REGION Network 13: DB60 DBX2.0 = FS332 No Flow
   // GCU_ALARM_WORD_02_BIT_0
   RUNG wire#powerrail
      Contact( "300_AUT_SEQ_TMRS_DB"."FS332 Delay".Q )
      { S7_Templates := "SrcType := Int" } GE_Contact(in1 := "100_GCU_AUTO_SEQ_DB".CRNT_STEP, in2 := 60)
      { S7_Templates := "SrcType := Int" } LE_Contact(in1 := "100_GCU_AUTO_SEQ_DB".CRNT_STEP, in2 := 560)
      S_Coil( %DB60.DBX2.0 )
   END_RUNG
   // the same network as SCL:
   IF "300_AUT_SEQ_TMRS_DB"."FS332 Delay".Q AND ("100_GCU_AUTO_SEQ_DB".CRNT_STEP >= 60) AND ("100_GCU_AUTO_SEQ_DB".CRNT_STEP <= 560) THEN
       %DB60.DBX2.0 := TRUE;
   END_IF;
END_REGION

REGION Network 14: DB60 DBX2.1 = PIT348 LOLO
   // GCU_ALARM_WORD_02_BIT_1      changed to 60 to 120 for test
   RUNG wire#powerrail
      { S7_Templates := "SrcType := Int" } GE_Contact(in1 := "100_GCU_AUTO_SEQ_DB".CRNT_STEP, in2 := 140)
      { S7_Templates := "SrcType := Int" } LT_Contact(in1 := "100_GCU_AUTO_SEQ_DB".CRNT_STEP, in2 := 540)
      Contact( "PIT348_ALM_ANALOG_DB73"."ALARM LL" )
      I_Contact( "10_DI_DATA"."FS_332 FLW_OK" )
      S_Coil( %DB60.DBX2.1 )
   END_RUNG
   // the same network as SCL:
   IF ("100_GCU_AUTO_SEQ_DB".CRNT_STEP >= 140) AND ("100_GCU_AUTO_SEQ_DB".CRNT_STEP < 540) AND "PIT348_ALM_ANALOG_DB73"."ALARM LL" AND NOT "10_DI_DATA"."FS_332 FLW_OK" THEN
       %DB60.DBX2.1 := TRUE;
   END_IF;
END_REGION

REGION Network 15: DB60 DBX2.2 = PIT348 HIHI
   // GCU_ALARM_WORD_02_BIT_2
   RUNG wire#powerrail
      Contact( "PIT348_ALM_ANALOG_DB73"."ALARM HH" )
      I_Contact( "10_DI_DATA"."FS_332 FLW_OK" )
      S_Coil( %DB60.DBX2.2 )
   END_RUNG
   // the same network as SCL:
   IF "PIT348_ALM_ANALOG_DB73"."ALARM HH" AND NOT "10_DI_DATA"."FS_332 FLW_OK" THEN
       %DB60.DBX2.2 := TRUE;
   END_IF;
END_REGION

REGION Network 16: DB60 DBX2.3 = FS350 Low Flow
   // GCU_ALARM_WORD_02_BIT_3
   RUNG wire#powerrail
      Contact( "TIT406_ALM_ANALOG_DB74".Error_present )
      Contact( "TIT408_ALM_ANALOG_DB75".Error_present )
      I_Contact( "10_DI_DATA".FS_350_FLW_OK )
      S_Coil( %DB60.DBX2.3 )
   END_RUNG
   // the same network as SCL:
   IF "TIT406_ALM_ANALOG_DB74".Error_present AND "TIT408_ALM_ANALOG_DB75".Error_present AND NOT "10_DI_DATA".FS_350_FLW_OK THEN
       %DB60.DBX2.3 := TRUE;
   END_IF;
END_REGION

REGION Network 17: DB60 DBX2.5 = TT002 HIHI
   // GCU_ALARM_WORD_02_BIT_5
   RUNG wire#powerrail
      Contact( "TT002_ALM_ANALOG_DB76"."ALARM HH" )
      S_Coil( %DB60.DBX2.5 )
   END_RUNG
   // the same network as SCL:
   IF "TT002_ALM_ANALOG_DB76"."ALARM HH" THEN %DB60.DBX2.5 := TRUE; END_IF;
END_REGION

REGION Network 18: DB60 DBX2.6 = PT002 HIHI
   // GCU_ALARM_WORD_02_BIT_6
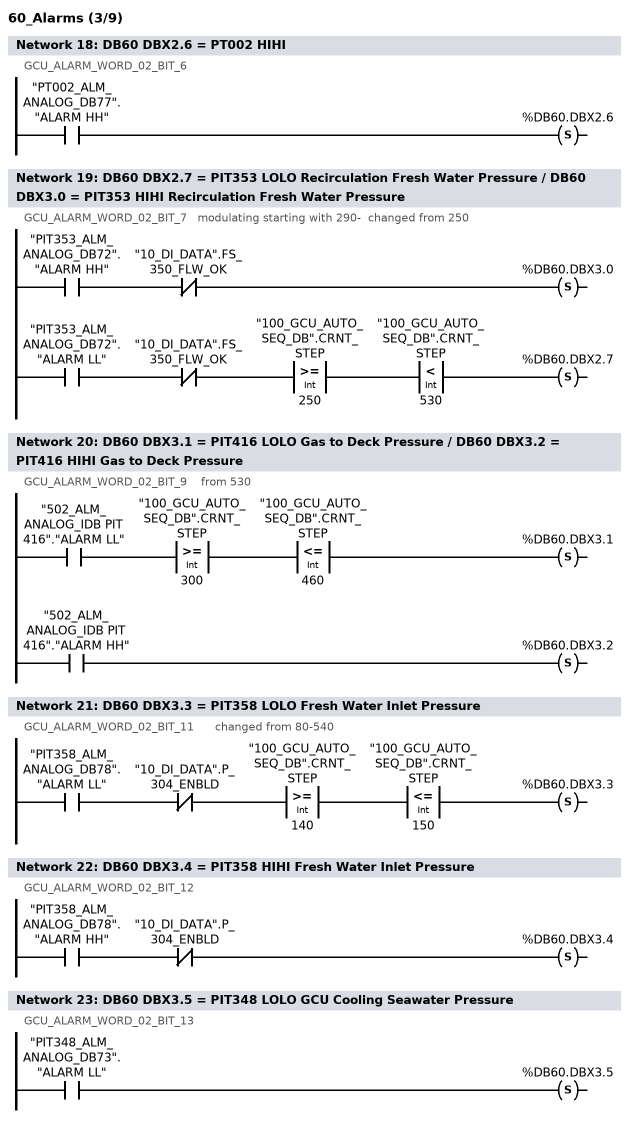
   RUNG wire#powerrail
      Contact( "PT002_ALM_ANALOG_DB77"."ALARM HH" )
      S_Coil( %DB60.DBX2.6 )
   END_RUNG
   // the same network as SCL:
   IF "PT002_ALM_ANALOG_DB77"."ALARM HH" THEN %DB60.DBX2.6 := TRUE; END_IF;
END_REGION

REGION Network 19: DB60 DBX2.7 = PIT353 LOLO Recirculation Fresh Water Pressure / DB60 DBX3.0 = PIT353 HIHI Recirculation Fresh Water Pressure
   // GCU_ALARM_WORD_02_BIT_7   modulating starting with 290-  changed from 250
   RUNG wire#powerrail
      Contact( "PIT353_ALM_ANALOG_DB72"."ALARM HH" )
      I_Contact( "10_DI_DATA".FS_350_FLW_OK )
      S_Coil( %DB60.DBX3.0 )
   END_RUNG
   RUNG wire#powerrail
      Contact( "PIT353_ALM_ANALOG_DB72"."ALARM LL" )
      I_Contact( "10_DI_DATA".FS_350_FLW_OK )
      { S7_Templates := "SrcType := Int" } GE_Contact(in1 := "100_GCU_AUTO_SEQ_DB".CRNT_STEP, in2 := 250)
      { S7_Templates := "SrcType := Int" } LT_Contact(in1 := "100_GCU_AUTO_SEQ_DB".CRNT_STEP, in2 := 530)
      S_Coil( %DB60.DBX2.7 )
   END_RUNG
   // the same network as SCL:
   IF "PIT353_ALM_ANALOG_DB72"."ALARM HH" AND NOT "10_DI_DATA".FS_350_FLW_OK THEN
       %DB60.DBX3.0 := TRUE;
   END_IF;
   IF "PIT353_ALM_ANALOG_DB72"."ALARM LL" AND NOT "10_DI_DATA".FS_350_FLW_OK AND ("100_GCU_AUTO_SEQ_DB".CRNT_STEP >= 250) AND ("100_GCU_AUTO_SEQ_DB".CRNT_STEP < 530) THEN
       %DB60.DBX2.7 := TRUE;
   END_IF;
END_REGION

REGION Network 20: DB60 DBX3.1 = PIT416 LOLO Gas to Deck Pressure / DB60 DBX3.2 = PIT416 HIHI Gas to Deck Pressure
   // GCU_ALARM_WORD_02_BIT_9    from 530
   RUNG wire#powerrail
      Contact( "502_ALM_ANALOG_IDB PIT 416"."ALARM LL" )
      { S7_Templates := "SrcType := Int" } GE_Contact(in1 := "100_GCU_AUTO_SEQ_DB".CRNT_STEP, in2 := 300)
      { S7_Templates := "SrcType := Int" } LE_Contact(in1 := "100_GCU_AUTO_SEQ_DB".CRNT_STEP, in2 := 460)
      S_Coil( %DB60.DBX3.1 )
   END_RUNG
   RUNG wire#powerrail
      Contact( "502_ALM_ANALOG_IDB PIT 416"."ALARM HH" )
      S_Coil( %DB60.DBX3.2 )
   END_RUNG
   // the same network as SCL:
   IF "502_ALM_ANALOG_IDB PIT 416"."ALARM LL" AND ("100_GCU_AUTO_SEQ_DB".CRNT_STEP >= 300) AND ("100_GCU_AUTO_SEQ_DB".CRNT_STEP <= 460) THEN
       %DB60.DBX3.1 := TRUE;
   END_IF;
   IF "502_ALM_ANALOG_IDB PIT 416"."ALARM HH" THEN %DB60.DBX3.2 := TRUE; END_IF;
END_REGION

REGION Network 21: DB60 DBX3.3 = PIT358 LOLO Fresh Water Inlet Pressure
   // GCU_ALARM_WORD_02_BIT_11      changed from 80-540
   RUNG wire#powerrail
      Contact( "PIT358_ALM_ANALOG_DB78"."ALARM LL" )
      I_Contact( "10_DI_DATA".P_304_ENBLD )
      { S7_Templates := "SrcType := Int" } GE_Contact(in1 := "100_GCU_AUTO_SEQ_DB".CRNT_STEP, in2 := 140)
      { S7_Templates := "SrcType := Int" } LE_Contact(in1 := "100_GCU_AUTO_SEQ_DB".CRNT_STEP, in2 := 150)
      S_Coil( %DB60.DBX3.3 )
   END_RUNG
   // the same network as SCL:
   IF "PIT358_ALM_ANALOG_DB78"."ALARM LL" AND NOT "10_DI_DATA".P_304_ENBLD AND ("100_GCU_AUTO_SEQ_DB".CRNT_STEP >= 140) AND ("100_GCU_AUTO_SEQ_DB".CRNT_STEP <= 150) THEN
       %DB60.DBX3.3 := TRUE;
   END_IF;
END_REGION

REGION Network 22: DB60 DBX3.4 = PIT358 HIHI Fresh Water Inlet Pressure
   // GCU_ALARM_WORD_02_BIT_12
   RUNG wire#powerrail
      Contact( "PIT358_ALM_ANALOG_DB78"."ALARM HH" )
      I_Contact( "10_DI_DATA".P_304_ENBLD )
      S_Coil( %DB60.DBX3.4 )
   END_RUNG
   // the same network as SCL:
   IF "PIT358_ALM_ANALOG_DB78"."ALARM HH" AND NOT "10_DI_DATA".P_304_ENBLD THEN %DB60.DBX3.4 := TRUE; END_IF;
END_REGION

REGION Network 23: DB60 DBX3.5 = PIT348 LOLO GCU Cooling Seawater Pressure
   // GCU_ALARM_WORD_02_BIT_13
   RUNG wire#powerrail
      Contact( "PIT348_ALM_ANALOG_DB73"."ALARM LL" )
      S_Coil( %DB60.DBX3.5 )
   END_RUNG
   // the same network as SCL:
   IF "PIT348_ALM_ANALOG_DB73"."ALARM LL" THEN %DB60.DBX3.5 := TRUE; END_IF;
END_REGION

REGION Network 24: DB60 DBX3.6 = PIT348 HIHI GCU Cooling Seawater Pressure
   // GCU_ALARM_WORD_02_BIT_14
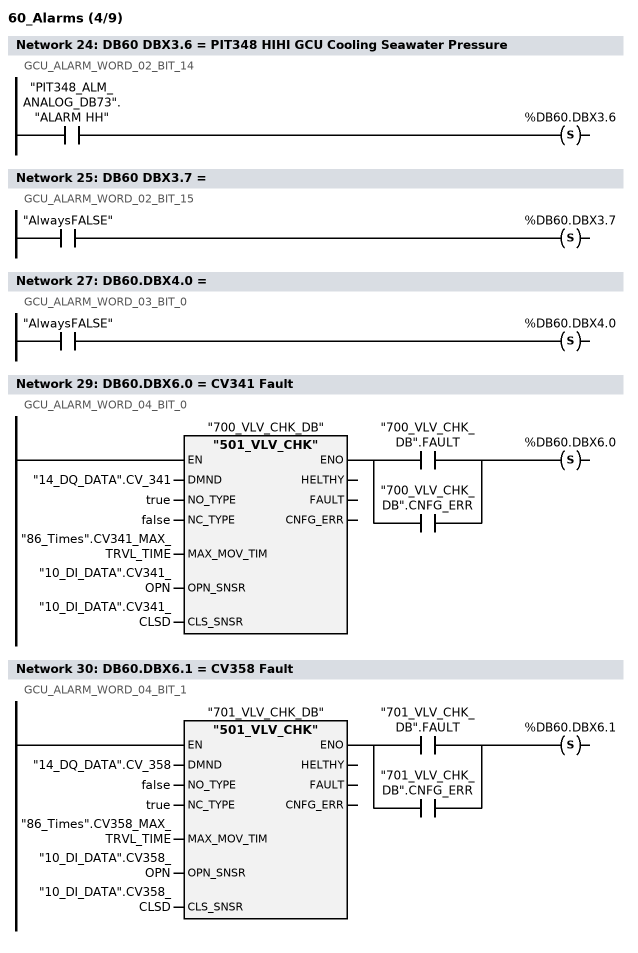
   RUNG wire#powerrail
      Contact( "PIT348_ALM_ANALOG_DB73"."ALARM HH" )
      S_Coil( %DB60.DBX3.6 )
   END_RUNG
   // the same network as SCL:
   IF "PIT348_ALM_ANALOG_DB73"."ALARM HH" THEN %DB60.DBX3.6 := TRUE; END_IF;
END_REGION

REGION Network 25: DB60 DBX3.7 =
   // GCU_ALARM_WORD_02_BIT_15
   RUNG wire#powerrail
      Contact( "AlwaysFALSE" )
      S_Coil( %DB60.DBX3.7 )
   END_RUNG
   // the same network as SCL:
   IF "AlwaysFALSE" THEN %DB60.DBX3.7 := TRUE; END_IF;
END_REGION

REGION Network 27: DB60.DBX4.0 =
   // GCU_ALARM_WORD_03_BIT_0
   RUNG wire#powerrail
      Contact( "AlwaysFALSE" )
      S_Coil( %DB60.DBX4.0 )
   END_RUNG
   // the same network as SCL:
   IF "AlwaysFALSE" THEN %DB60.DBX4.0 := TRUE; END_IF;
END_REGION

REGION Network 29: DB60.DBX6.0 = CV341 Fault
   // GCU_ALARM_WORD_04_BIT_0
   RUNG wire#powerrail
      "700_VLV_CHK_DB"(DMND := "14_DQ_DATA".CV_341, NO_TYPE := true, NC_TYPE := false, MAX_MOV_TIM := "86_Times".CV341_MAX_TRVL_TIME, OPN_SNSR := "10_DI_DATA".CV341_OPN, CLS_SNSR := "10_DI_DATA".CV341_CLSD, HELTHY =>, FAULT =>, CNFG_ERR =>)
      wire#w1
      Contact( "700_VLV_CHK_DB".FAULT )
      wire#w2
      S_Coil( %DB60.DBX6.0 )
   END_RUNG
   RUNG wire#w1
      Contact( "700_VLV_CHK_DB".CNFG_ERR )
   END_RUNG wire#w2
   // the same network as SCL:
   "700_VLV_CHK_DB"(DMND := "14_DQ_DATA".CV_341,   // "501_VLV_CHK"
                    NO_TYPE := true,
                    NC_TYPE := false,
                    MAX_MOV_TIM := "86_Times".CV341_MAX_TRVL_TIME,
                    OPN_SNSR := "10_DI_DATA".CV341_OPN,
                    CLS_SNSR := "10_DI_DATA".CV341_CLSD,
                    ENO => #_w1);
   IF #_w1 AND ("700_VLV_CHK_DB".FAULT OR "700_VLV_CHK_DB".CNFG_ERR) THEN %DB60.DBX6.0 := TRUE; END_IF;
END_REGION

REGION Network 30: DB60.DBX6.1 = CV358 Fault
   // GCU_ALARM_WORD_04_BIT_1
   RUNG wire#powerrail
      "701_VLV_CHK_DB"(DMND := "14_DQ_DATA".CV_358, NO_TYPE := false, NC_TYPE := true, MAX_MOV_TIM := "86_Times".CV358_MAX_TRVL_TIME, OPN_SNSR := "10_DI_DATA".CV358_OPN, CLS_SNSR := "10_DI_DATA".CV358_CLSD, HELTHY =>, FAULT =>, CNFG_ERR =>)
      wire#w1
      Contact( "701_VLV_CHK_DB".FAULT )
      wire#w2
      S_Coil( %DB60.DBX6.1 )
   END_RUNG
   RUNG wire#w1
      Contact( "701_VLV_CHK_DB".CNFG_ERR )
   END_RUNG wire#w2
   // the same network as SCL:
   "701_VLV_CHK_DB"(DMND := "14_DQ_DATA".CV_358,   // "501_VLV_CHK"
                    NO_TYPE := false,
                    NC_TYPE := true,
                    MAX_MOV_TIM := "86_Times".CV358_MAX_TRVL_TIME,
                    OPN_SNSR := "10_DI_DATA".CV358_OPN,
                    CLS_SNSR := "10_DI_DATA".CV358_CLSD,
                    ENO => #_w1);
   IF #_w1 AND ("701_VLV_CHK_DB".FAULT OR "701_VLV_CHK_DB".CNFG_ERR) THEN %DB60.DBX6.1 := TRUE; END_IF;
END_REGION

REGION Network 31: DB60.DBX6.2 = CV406 Fault
   // GCU_ALARM_WORD_04_BIT_2
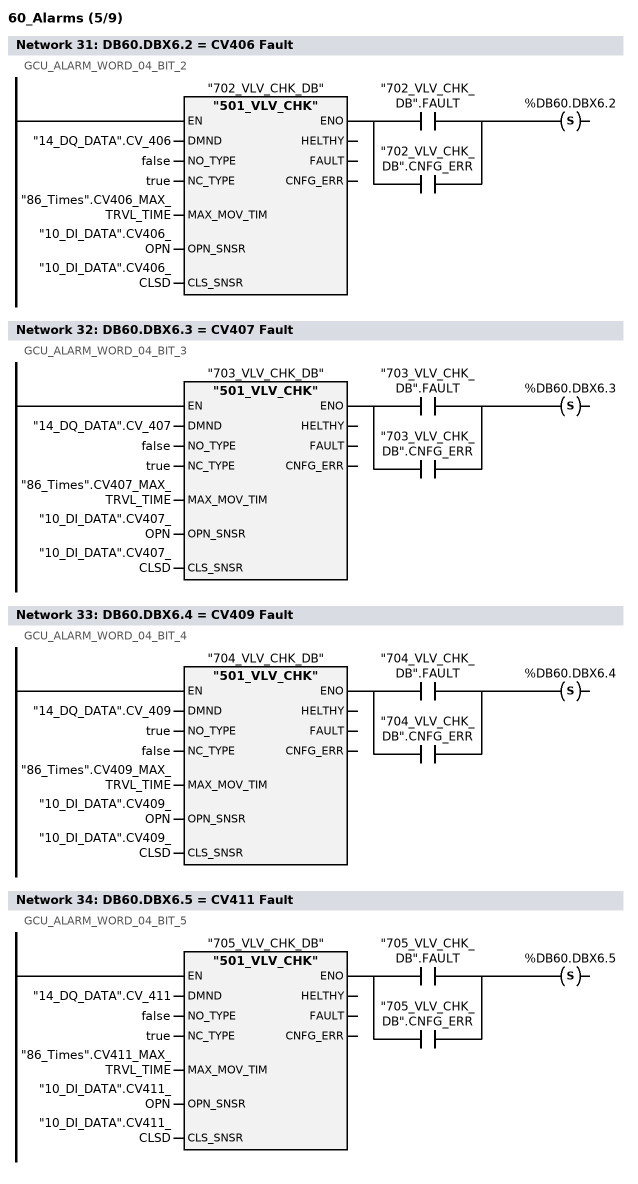
   RUNG wire#powerrail
      "702_VLV_CHK_DB"(DMND := "14_DQ_DATA".CV_406, NO_TYPE := false, NC_TYPE := true, MAX_MOV_TIM := "86_Times".CV406_MAX_TRVL_TIME, OPN_SNSR := "10_DI_DATA".CV406_OPN, CLS_SNSR := "10_DI_DATA".CV406_CLSD, HELTHY =>, FAULT =>, CNFG_ERR =>)
      wire#w1
      Contact( "702_VLV_CHK_DB".FAULT )
      wire#w2
      S_Coil( %DB60.DBX6.2 )
   END_RUNG
   RUNG wire#w1
      Contact( "702_VLV_CHK_DB".CNFG_ERR )
   END_RUNG wire#w2
   // the same network as SCL:
   "702_VLV_CHK_DB"(DMND := "14_DQ_DATA".CV_406,   // "501_VLV_CHK"
                    NO_TYPE := false,
                    NC_TYPE := true,
                    MAX_MOV_TIM := "86_Times".CV406_MAX_TRVL_TIME,
                    OPN_SNSR := "10_DI_DATA".CV406_OPN,
                    CLS_SNSR := "10_DI_DATA".CV406_CLSD,
                    ENO => #_w1);
   IF #_w1 AND ("702_VLV_CHK_DB".FAULT OR "702_VLV_CHK_DB".CNFG_ERR) THEN %DB60.DBX6.2 := TRUE; END_IF;
END_REGION

REGION Network 32: DB60.DBX6.3 = CV407 Fault
   // GCU_ALARM_WORD_04_BIT_3
   RUNG wire#powerrail
      "703_VLV_CHK_DB"(DMND := "14_DQ_DATA".CV_407, NO_TYPE := false, NC_TYPE := true, MAX_MOV_TIM := "86_Times".CV407_MAX_TRVL_TIME, OPN_SNSR := "10_DI_DATA".CV407_OPN, CLS_SNSR := "10_DI_DATA".CV407_CLSD, HELTHY =>, FAULT =>, CNFG_ERR =>)
      wire#w1
      Contact( "703_VLV_CHK_DB".FAULT )
      wire#w2
      S_Coil( %DB60.DBX6.3 )
   END_RUNG
   RUNG wire#w1
      Contact( "703_VLV_CHK_DB".CNFG_ERR )
   END_RUNG wire#w2
   // the same network as SCL:
   "703_VLV_CHK_DB"(DMND := "14_DQ_DATA".CV_407,   // "501_VLV_CHK"
                    NO_TYPE := false,
                    NC_TYPE := true,
                    MAX_MOV_TIM := "86_Times".CV407_MAX_TRVL_TIME,
                    OPN_SNSR := "10_DI_DATA".CV407_OPN,
                    CLS_SNSR := "10_DI_DATA".CV407_CLSD,
                    ENO => #_w1);
   IF #_w1 AND ("703_VLV_CHK_DB".FAULT OR "703_VLV_CHK_DB".CNFG_ERR) THEN %DB60.DBX6.3 := TRUE; END_IF;
END_REGION

REGION Network 33: DB60.DBX6.4 = CV409 Fault
   // GCU_ALARM_WORD_04_BIT_4
   RUNG wire#powerrail
      "704_VLV_CHK_DB"(DMND := "14_DQ_DATA".CV_409, NO_TYPE := true, NC_TYPE := false, MAX_MOV_TIM := "86_Times".CV409_MAX_TRVL_TIME, OPN_SNSR := "10_DI_DATA".CV409_OPN, CLS_SNSR := "10_DI_DATA".CV409_CLSD, HELTHY =>, FAULT =>, CNFG_ERR =>)
      wire#w1
      Contact( "704_VLV_CHK_DB".FAULT )
      wire#w2
      S_Coil( %DB60.DBX6.4 )
   END_RUNG
   RUNG wire#w1
      Contact( "704_VLV_CHK_DB".CNFG_ERR )
   END_RUNG wire#w2
   // the same network as SCL:
   "704_VLV_CHK_DB"(DMND := "14_DQ_DATA".CV_409,   // "501_VLV_CHK"
                    NO_TYPE := true,
                    NC_TYPE := false,
                    MAX_MOV_TIM := "86_Times".CV409_MAX_TRVL_TIME,
                    OPN_SNSR := "10_DI_DATA".CV409_OPN,
                    CLS_SNSR := "10_DI_DATA".CV409_CLSD,
                    ENO => #_w1);
   IF #_w1 AND ("704_VLV_CHK_DB".FAULT OR "704_VLV_CHK_DB".CNFG_ERR) THEN %DB60.DBX6.4 := TRUE; END_IF;
END_REGION

REGION Network 34: DB60.DBX6.5 = CV411 Fault
   // GCU_ALARM_WORD_04_BIT_5
   RUNG wire#powerrail
      "705_VLV_CHK_DB"(DMND := "14_DQ_DATA".CV_411, NO_TYPE := false, NC_TYPE := true, MAX_MOV_TIM := "86_Times".CV411_MAX_TRVL_TIME, OPN_SNSR := "10_DI_DATA".CV411_OPN, CLS_SNSR := "10_DI_DATA".CV411_CLSD, HELTHY =>, FAULT =>, CNFG_ERR =>)
      wire#w1
      Contact( "705_VLV_CHK_DB".FAULT )
      wire#w2
      S_Coil( %DB60.DBX6.5 )
   END_RUNG
   RUNG wire#w1
      Contact( "705_VLV_CHK_DB".CNFG_ERR )
   END_RUNG wire#w2
   // the same network as SCL:
   "705_VLV_CHK_DB"(DMND := "14_DQ_DATA".CV_411,   // "501_VLV_CHK"
                    NO_TYPE := false,
                    NC_TYPE := true,
                    MAX_MOV_TIM := "86_Times".CV411_MAX_TRVL_TIME,
                    OPN_SNSR := "10_DI_DATA".CV411_OPN,
                    CLS_SNSR := "10_DI_DATA".CV411_CLSD,
                    ENO => #_w1);
   IF #_w1 AND ("705_VLV_CHK_DB".FAULT OR "705_VLV_CHK_DB".CNFG_ERR) THEN %DB60.DBX6.5 := TRUE; END_IF;
END_REGION

REGION Network 35: DB60.DBX6.6 = CV441 Fault
   // GCU_ALARM_WORD_04_BIT_6
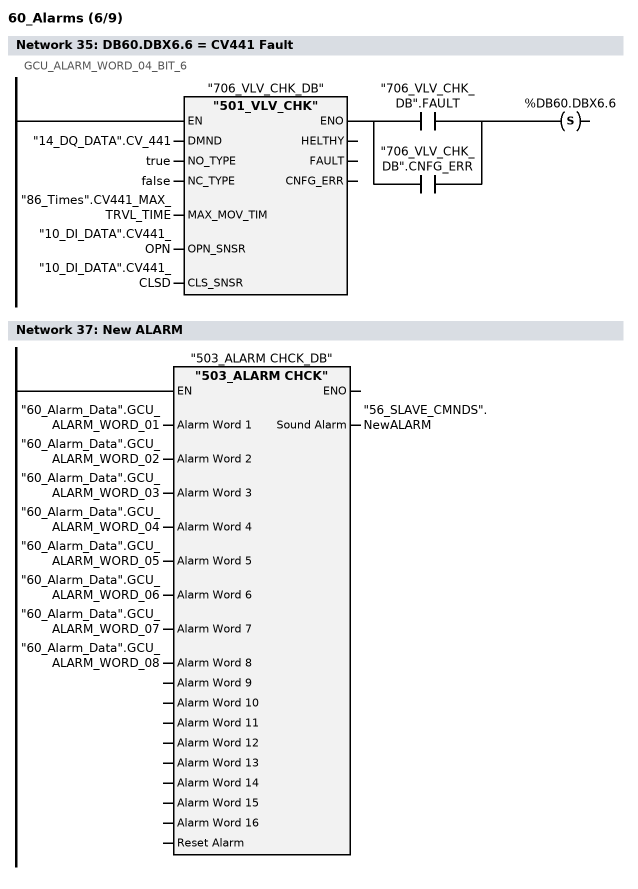
   RUNG wire#powerrail
      "706_VLV_CHK_DB"(DMND := "14_DQ_DATA".CV_441, NO_TYPE := true, NC_TYPE := false, MAX_MOV_TIM := "86_Times".CV441_MAX_TRVL_TIME, OPN_SNSR := "10_DI_DATA".CV441_OPN, CLS_SNSR := "10_DI_DATA".CV441_CLSD, HELTHY =>, FAULT =>, CNFG_ERR =>)
      wire#w1
      Contact( "706_VLV_CHK_DB".FAULT )
      wire#w2
      S_Coil( %DB60.DBX6.6 )
   END_RUNG
   RUNG wire#w1
      Contact( "706_VLV_CHK_DB".CNFG_ERR )
   END_RUNG wire#w2
   // the same network as SCL:
   "706_VLV_CHK_DB"(DMND := "14_DQ_DATA".CV_441,   // "501_VLV_CHK"
                    NO_TYPE := true,
                    NC_TYPE := false,
                    MAX_MOV_TIM := "86_Times".CV441_MAX_TRVL_TIME,
                    OPN_SNSR := "10_DI_DATA".CV441_OPN,
                    CLS_SNSR := "10_DI_DATA".CV441_CLSD,
                    ENO => #_w1);
   IF #_w1 AND ("706_VLV_CHK_DB".FAULT OR "706_VLV_CHK_DB".CNFG_ERR) THEN %DB60.DBX6.6 := TRUE; END_IF;
END_REGION

REGION Network 37: New ALARM
   RUNG wire#powerrail
      "503_ALARM CHCK_DB"("Alarm Word 1" := "60_Alarm_Data".GCU_ALARM_WORD_01, "Alarm Word 2" := "60_Alarm_Data".GCU_ALARM_WORD_02, "Alarm Word 3" := "60_Alarm_Data".GCU_ALARM_WORD_03, "Alarm Word 4" := "60_Alarm_Data".GCU_ALARM_WORD_04, "Alarm Word 5" := "60_Alarm_Data".GCU_ALARM_WORD_05, "Alarm Word 6" := "60_Alarm_Data".GCU_ALARM_WORD_06, "Alarm Word 7" := "60_Alarm_Data".GCU_ALARM_WORD_07, "Alarm Word 8" := "60_Alarm_Data".GCU_ALARM_WORD_08, "Alarm Word 9" :=, "Alarm Word 10" :=, "Alarm Word 11" :=, "Alarm Word 12" :=, "Alarm Word 13" :=, "Alarm Word 14" :=, "Alarm Word 15" :=, "Alarm Word 16" :=, "Reset Alarm" :=, "Sound Alarm" => "56_SLAVE_CMNDS".NewALARM)
   END_RUNG
   // the same network as SCL:
   "503_ALARM CHCK_DB"("Alarm Word 1" := "60_Alarm_Data".GCU_ALARM_WORD_01,   // "503_ALARM CHCK"
                       "Alarm Word 2" := "60_Alarm_Data".GCU_ALARM_WORD_02,
                       "Alarm Word 3" := "60_Alarm_Data".GCU_ALARM_WORD_03,
                       "Alarm Word 4" := "60_Alarm_Data".GCU_ALARM_WORD_04,
                       "Alarm Word 5" := "60_Alarm_Data".GCU_ALARM_WORD_05,
                       "Alarm Word 6" := "60_Alarm_Data".GCU_ALARM_WORD_06,
                       "Alarm Word 7" := "60_Alarm_Data".GCU_ALARM_WORD_07,
                       "Alarm Word 8" := "60_Alarm_Data".GCU_ALARM_WORD_08,
                       "Sound Alarm" => "56_SLAVE_CMNDS".NewALARM);
END_REGION

REGION Network 38: Alarm Present
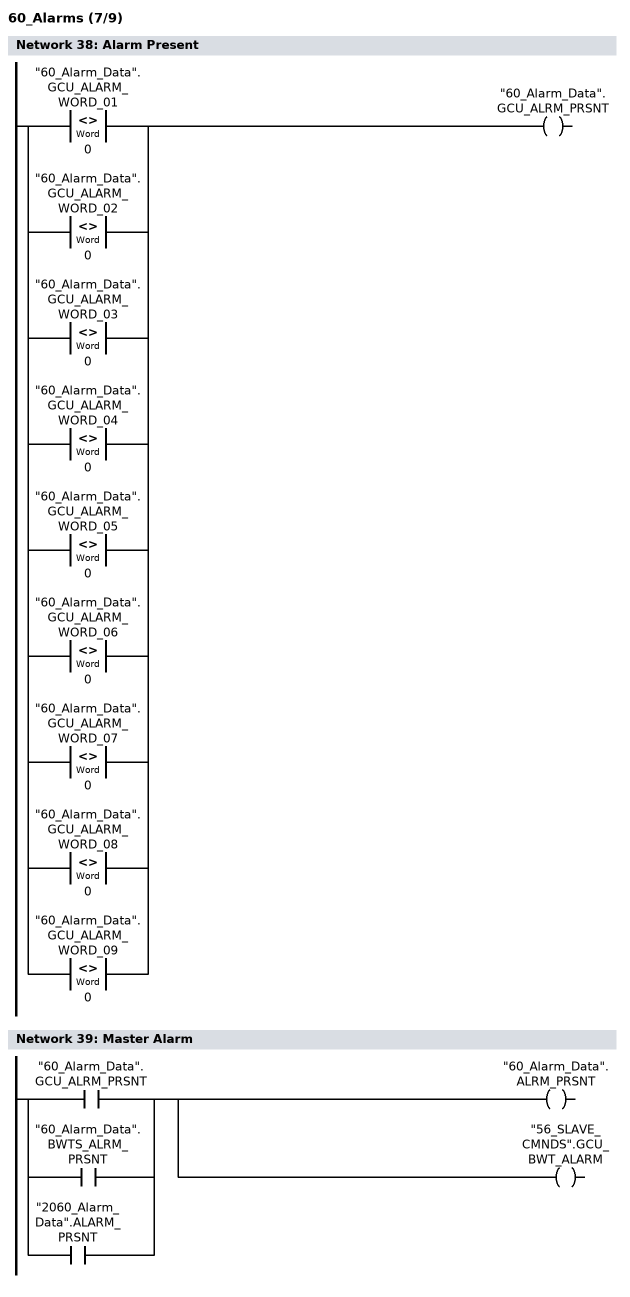
   RUNG wire#powerrail
      { S7_Templates := "SrcType := Word" } NE_Contact(in1 := "60_Alarm_Data".GCU_ALARM_WORD_01, in2 := 0)
      wire#w1
      Coil( "60_Alarm_Data".GCU_ALRM_PRSNT )
   END_RUNG
   RUNG wire#powerrail
      { S7_Templates := "SrcType := Word" } NE_Contact(in1 := "60_Alarm_Data".GCU_ALARM_WORD_02, in2 := 0)
   END_RUNG wire#w1
   RUNG wire#powerrail
      { S7_Templates := "SrcType := Word" } NE_Contact(in1 := "60_Alarm_Data".GCU_ALARM_WORD_03, in2 := 0)
   END_RUNG wire#w1
   RUNG wire#powerrail
      { S7_Templates := "SrcType := Word" } NE_Contact(in1 := "60_Alarm_Data".GCU_ALARM_WORD_04, in2 := 0)
   END_RUNG wire#w1
   RUNG wire#powerrail
      { S7_Templates := "SrcType := Word" } NE_Contact(in1 := "60_Alarm_Data".GCU_ALARM_WORD_05, in2 := 0)
   END_RUNG wire#w1
   RUNG wire#powerrail
      { S7_Templates := "SrcType := Word" } NE_Contact(in1 := "60_Alarm_Data".GCU_ALARM_WORD_06, in2 := 0)
   END_RUNG wire#w1
   RUNG wire#powerrail
      { S7_Templates := "SrcType := Word" } NE_Contact(in1 := "60_Alarm_Data".GCU_ALARM_WORD_07, in2 := 0)
   END_RUNG wire#w1
   RUNG wire#powerrail
      { S7_Templates := "SrcType := Word" } NE_Contact(in1 := "60_Alarm_Data".GCU_ALARM_WORD_08, in2 := 0)
   END_RUNG wire#w1
   RUNG wire#powerrail
      { S7_Templates := "SrcType := Word" } NE_Contact(in1 := "60_Alarm_Data".GCU_ALARM_WORD_09, in2 := 0)
   END_RUNG wire#w1
   // the same network as SCL:
   "60_Alarm_Data".GCU_ALRM_PRSNT := ("60_Alarm_Data".GCU_ALARM_WORD_01 <> 0) OR ("60_Alarm_Data".GCU_ALARM_WORD_02 <> 0) OR ("60_Alarm_Data".GCU_ALARM_WORD_03 <> 0) OR ("60_Alarm_Data".GCU_ALARM_WORD_04 <> 0) OR ("60_Alarm_Data".GCU_ALARM_WORD_05 <> 0) OR ("60_Alarm_Data".GCU_ALARM_WORD_06 <> 0) OR ("60_Alarm_Data".GCU_ALARM_WORD_07 <> 0) OR ("60_Alarm_Data".GCU_ALARM_WORD_08 <> 0) OR ("60_Alarm_Data".GCU_ALARM_WORD_09 <> 0);
END_REGION

REGION Network 39: Master Alarm
   RUNG wire#powerrail
      Contact( "60_Alarm_Data".GCU_ALRM_PRSNT )
      wire#w1
      Coil( "60_Alarm_Data".ALRM_PRSNT )
   END_RUNG
   RUNG wire#powerrail
      Contact( "60_Alarm_Data".BWTS_ALRM_PRSNT )
   END_RUNG wire#w1
   RUNG wire#powerrail
      Contact( "2060_Alarm_Data".ALARM_PRSNT )
   END_RUNG wire#w1
   RUNG wire#w1
      Coil( "56_SLAVE_CMNDS".GCU_BWT_ALARM )
   END_RUNG
   // the same network as SCL:
   "60_Alarm_Data".ALRM_PRSNT := "60_Alarm_Data".GCU_ALRM_PRSNT OR "60_Alarm_Data".BWTS_ALRM_PRSNT OR "2060_Alarm_Data".ALARM_PRSNT;
   "56_SLAVE_CMNDS".GCU_BWT_ALARM := "60_Alarm_Data".ALRM_PRSNT;
END_REGION

REGION Network 40: Alarm reset
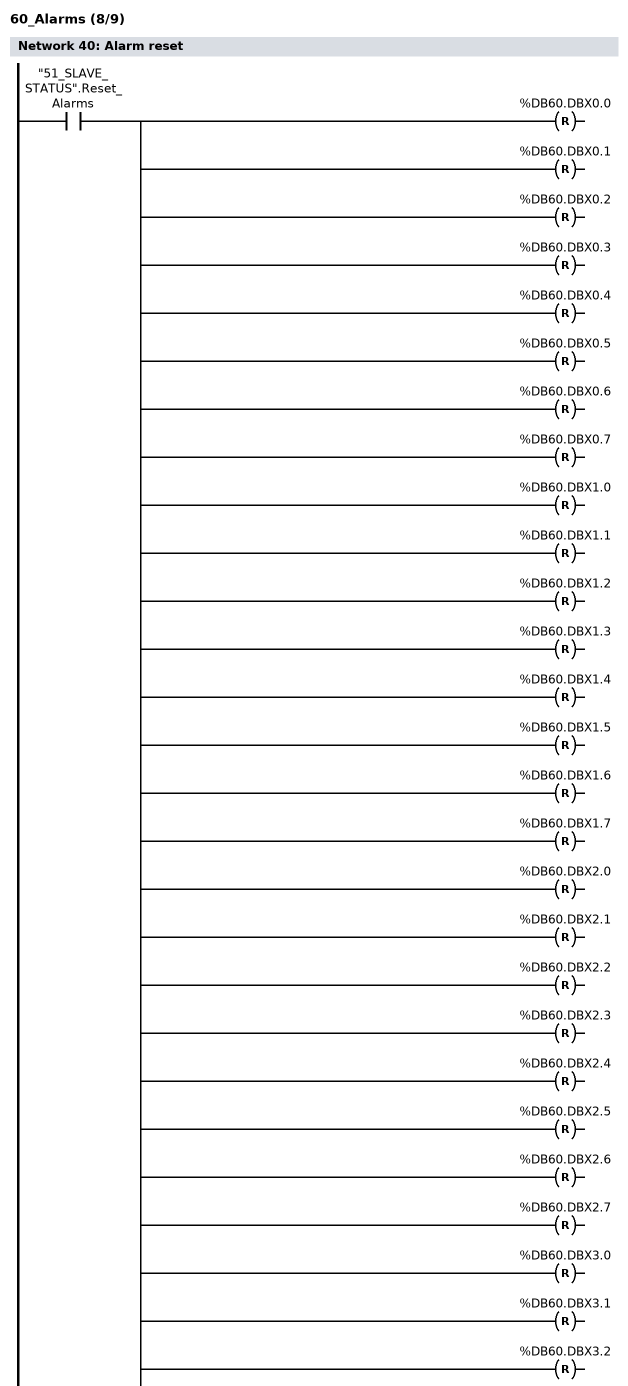
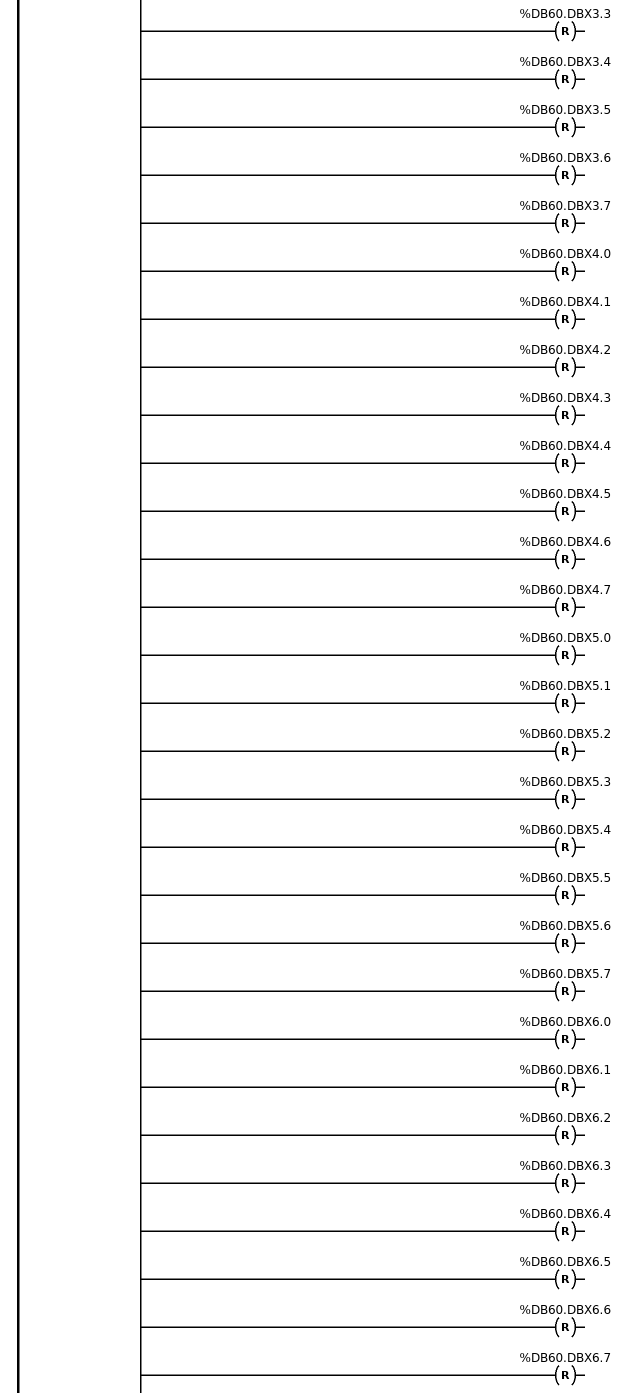
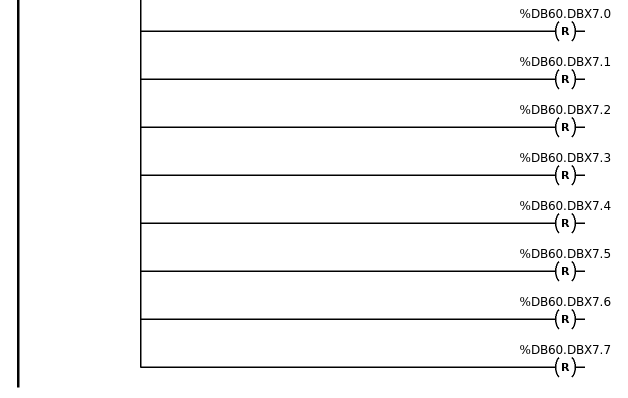
   RUNG wire#powerrail
      Contact( "51_SLAVE_STATUS".Reset_Alarms )
      wire#w1
      R_Coil( %DB60.DBX0.0 )
   END_RUNG
   RUNG wire#w1
      R_Coil( %DB60.DBX0.1 )
   END_RUNG
   RUNG wire#w1
      R_Coil( %DB60.DBX0.2 )
   END_RUNG
   RUNG wire#w1
      R_Coil( %DB60.DBX0.3 )
   END_RUNG
   RUNG wire#w1
      R_Coil( %DB60.DBX0.4 )
   END_RUNG
   RUNG wire#w1
      R_Coil( %DB60.DBX0.5 )
   END_RUNG
   RUNG wire#w1
      R_Coil( %DB60.DBX0.6 )
   END_RUNG
   RUNG wire#w1
      R_Coil( %DB60.DBX0.7 )
   END_RUNG
   RUNG wire#w1
      R_Coil( %DB60.DBX1.0 )
   END_RUNG
   RUNG wire#w1
      R_Coil( %DB60.DBX1.1 )
   END_RUNG
   RUNG wire#w1
      R_Coil( %DB60.DBX1.2 )
   END_RUNG
   RUNG wire#w1
      R_Coil( %DB60.DBX1.3 )
   END_RUNG
   RUNG wire#w1
      R_Coil( %DB60.DBX1.4 )
   END_RUNG
   RUNG wire#w1
      R_Coil( %DB60.DBX1.5 )
   END_RUNG
   RUNG wire#w1
      R_Coil( %DB60.DBX1.6 )
   END_RUNG
   RUNG wire#w1
      R_Coil( %DB60.DBX1.7 )
   END_RUNG
   RUNG wire#w1
      R_Coil( %DB60.DBX2.0 )
   END_RUNG
   RUNG wire#w1
      R_Coil( %DB60.DBX2.1 )
   END_RUNG
   RUNG wire#w1
      R_Coil( %DB60.DBX2.2 )
   END_RUNG
   RUNG wire#w1
      R_Coil( %DB60.DBX2.3 )
   END_RUNG
   RUNG wire#w1
      R_Coil( %DB60.DBX2.4 )
   END_RUNG
   RUNG wire#w1
      R_Coil( %DB60.DBX2.5 )
   END_RUNG
   RUNG wire#w1
      R_Coil( %DB60.DBX2.6 )
   END_RUNG
   RUNG wire#w1
      R_Coil( %DB60.DBX2.7 )
   END_RUNG
   RUNG wire#w1
      R_Coil( %DB60.DBX3.0 )
   END_RUNG
   RUNG wire#w1
      R_Coil( %DB60.DBX3.1 )
   END_RUNG
   RUNG wire#w1
      R_Coil( %DB60.DBX3.2 )
   END_RUNG
   RUNG wire#w1
      R_Coil( %DB60.DBX3.3 )
   END_RUNG
   RUNG wire#w1
      R_Coil( %DB60.DBX3.4 )
   END_RUNG
   RUNG wire#w1
      R_Coil( %DB60.DBX3.5 )
   END_RUNG
   RUNG wire#w1
      R_Coil( %DB60.DBX3.6 )
   END_RUNG
   RUNG wire#w1
      R_Coil( %DB60.DBX3.7 )
   END_RUNG
   RUNG wire#w1
      R_Coil( %DB60.DBX4.0 )
   END_RUNG
   RUNG wire#w1
      R_Coil( %DB60.DBX4.1 )
   END_RUNG
   RUNG wire#w1
      R_Coil( %DB60.DBX4.2 )
   END_RUNG
   RUNG wire#w1
      R_Coil( %DB60.DBX4.3 )
   END_RUNG
   RUNG wire#w1
      R_Coil( %DB60.DBX4.4 )
   END_RUNG
   RUNG wire#w1
      R_Coil( %DB60.DBX4.5 )
   END_RUNG
   RUNG wire#w1
      R_Coil( %DB60.DBX4.6 )
   END_RUNG
   RUNG wire#w1
      R_Coil( %DB60.DBX4.7 )
   END_RUNG
   RUNG wire#w1
      R_Coil( %DB60.DBX5.0 )
   END_RUNG
   RUNG wire#w1
      R_Coil( %DB60.DBX5.1 )
   END_RUNG
   RUNG wire#w1
      R_Coil( %DB60.DBX5.2 )
   END_RUNG
   RUNG wire#w1
      R_Coil( %DB60.DBX5.3 )
   END_RUNG
   RUNG wire#w1
      R_Coil( %DB60.DBX5.4 )
   END_RUNG
   RUNG wire#w1
      R_Coil( %DB60.DBX5.5 )
   END_RUNG
   RUNG wire#w1
      R_Coil( %DB60.DBX5.6 )
   END_RUNG
   RUNG wire#w1
      R_Coil( %DB60.DBX5.7 )
   END_RUNG
   RUNG wire#w1
      R_Coil( %DB60.DBX6.0 )
   END_RUNG
   RUNG wire#w1
      R_Coil( %DB60.DBX6.1 )
   END_RUNG
   RUNG wire#w1
      R_Coil( %DB60.DBX6.2 )
   END_RUNG
   RUNG wire#w1
      R_Coil( %DB60.DBX6.3 )
   END_RUNG
   RUNG wire#w1
      R_Coil( %DB60.DBX6.4 )
   END_RUNG
   RUNG wire#w1
      R_Coil( %DB60.DBX6.5 )
   END_RUNG
   RUNG wire#w1
      R_Coil( %DB60.DBX6.6 )
   END_RUNG
   RUNG wire#w1
      R_Coil( %DB60.DBX6.7 )
   END_RUNG
   RUNG wire#w1
      R_Coil( %DB60.DBX7.0 )
   END_RUNG
   RUNG wire#w1
      R_Coil( %DB60.DBX7.1 )
   END_RUNG
   RUNG wire#w1
      R_Coil( %DB60.DBX7.2 )
   END_RUNG
   RUNG wire#w1
      R_Coil( %DB60.DBX7.3 )
   END_RUNG
   RUNG wire#w1
      R_Coil( %DB60.DBX7.4 )
   END_RUNG
   RUNG wire#w1
      R_Coil( %DB60.DBX7.5 )
   END_RUNG
   RUNG wire#w1
      R_Coil( %DB60.DBX7.6 )
   END_RUNG
   RUNG wire#w1
      R_Coil( %DB60.DBX7.7 )
   END_RUNG
   // the same network as SCL:
   IF "51_SLAVE_STATUS".Reset_Alarms THEN
       %DB60.DBX0.0 := FALSE;
       %DB60.DBX0.1 := FALSE;
       %DB60.DBX0.2 := FALSE;
       %DB60.DBX0.3 := FALSE;
       %DB60.DBX0.4 := FALSE;
       %DB60.DBX0.5 := FALSE;
       %DB60.DBX0.6 := FALSE;
       %DB60.DBX0.7 := FALSE;
       %DB60.DBX1.0 := FALSE;
       %DB60.DBX1.1 := FALSE;
       %DB60.DBX1.2 := FALSE;
       %DB60.DBX1.3 := FALSE;
       %DB60.DBX1.4 := FALSE;
       %DB60.DBX1.5 := FALSE;
       %DB60.DBX1.6 := FALSE;
       %DB60.DBX1.7 := FALSE;
       %DB60.DBX2.0 := FALSE;
       %DB60.DBX2.1 := FALSE;
       %DB60.DBX2.2 := FALSE;
       %DB60.DBX2.3 := FALSE;
       %DB60.DBX2.4 := FALSE;
       %DB60.DBX2.5 := FALSE;
       %DB60.DBX2.6 := FALSE;
       %DB60.DBX2.7 := FALSE;
       %DB60.DBX3.0 := FALSE;
       %DB60.DBX3.1 := FALSE;
       %DB60.DBX3.2 := FALSE;
       %DB60.DBX3.3 := FALSE;
       %DB60.DBX3.4 := FALSE;
       %DB60.DBX3.5 := FALSE;
       %DB60.DBX3.6 := FALSE;
       %DB60.DBX3.7 := FALSE;
       %DB60.DBX4.0 := FALSE;
       %DB60.DBX4.1 := FALSE;
       %DB60.DBX4.2 := FALSE;
       %DB60.DBX4.3 := FALSE;
       %DB60.DBX4.4 := FALSE;
       %DB60.DBX4.5 := FALSE;
       %DB60.DBX4.6 := FALSE;
       %DB60.DBX4.7 := FALSE;
       %DB60.DBX5.0 := FALSE;
       %DB60.DBX5.1 := FALSE;
       %DB60.DBX5.2 := FALSE;
       %DB60.DBX5.3 := FALSE;
       %DB60.DBX5.4 := FALSE;
       %DB60.DBX5.5 := FALSE;
       %DB60.DBX5.6 := FALSE;
       %DB60.DBX5.7 := FALSE;
       %DB60.DBX6.0 := FALSE;
       %DB60.DBX6.1 := FALSE;
       %DB60.DBX6.2 := FALSE;
       %DB60.DBX6.3 := FALSE;
       %DB60.DBX6.4 := FALSE;
       %DB60.DBX6.5 := FALSE;
       %DB60.DBX6.6 := FALSE;
       %DB60.DBX6.7 := FALSE;
       %DB60.DBX7.0 := FALSE;
       %DB60.DBX7.1 := FALSE;
       %DB60.DBX7.2 := FALSE;
       %DB60.DBX7.3 := FALSE;
       %DB60.DBX7.4 := FALSE;
       %DB60.DBX7.5 := FALSE;
       %DB60.DBX7.6 := FALSE;
       %DB60.DBX7.7 := FALSE;
   END_IF;
END_REGION

REGION Network 41: Step Set With Alarm
